text list "msjOp0": 20 'Alarma produs aparut anormal Confirmati prezenta ,integritatea si pozitia produs(planeitate , incadrarea in margini).'; 10 'Alarma detectie produs pierduta Verificati daca produsul mai exista in statie'; 11 'Alarma detectie produs pierduta Produsul exista dar nu e detectat. Reparati/ajustati senzorul de prezenta ssssssssssssssss,astfel incat sa detecteze produsul.'; 21 'Alarma produs aparut anormal Produsul nu a fost confirmat de operator Reparati senzorul ca sa nu mai indice prezenta produs'; 30 'Produsul nu a ajuns de la primul punct la al 2 lea Confirmati unde e de fapt produsul.'; 70 'Aduceti cilindru cccccccccccccc in pozitia xxxxxxxxxxxxxxx'; 72 'Deoarece a fost o alarma de griper confirmati prezenta ,integritatea si pozitia produs(planeitate , incadrarea in margini) in griper cccccccccccccc si lipsa lui de pe conveyor'; 73 'Deoarece a fost o alarma de griper confirmati prezenta ,integritatea si pozitia produs(planeitate , incadrarea in margini) pe palet si lipsa lui din griper cccccccccccccccccc'; 74 'Deoarece a fost o eroare de cilindru,confirmati ca liftul e sus si pachetul asezat pe el'; 71 ''; 22 'Alarma produs aparut anormal Produsul nu e asezat corect. Deschideti usa si plasati corect sau evacuati manual produsul,apoi validati'; 12 'Alarma detectie produs pierduta Produsul exista dar e prost asezat Deschideti usa si asezati sau eliminati produsul ,apoi confirmati.'; 31 'Produsul nu a ajuns de la primul punct la al 2 lea Produsul exista la destinatie dar nu e detectat.Deschideti usa si asezati produsul in dreptul senzorului ,sau reparati senzorul astfel incat sa detecteze produsul'; 32 'Produsul nu a ajuns de la primul punct la al 2 lea Produsul a ajuns la destinatie . Verificati prezenta,integritatea si pozitia lui si confirmati .'; 33 'Produsul nu a ajuns de la primul punct la al 2 lea Produsul a disparut din zona in mod necontrolat .Confirmati ca nici un produs nu se gaseste intre cele 2 posturi ,pentru a declara zona goala, si a putea accepta alte produse.'; 13 'Alarma detectie produs pierduta Detectia produsului a revenit Confirmati existenta si pozitia produs.'; 23 'Alarma produs aparut anormal Detectia produsului a disparut. Confirmati daca produsul mai exista'; 75 ''; 14 'Alarma detectie produs pierduta Produsul nu exista dar e detectat. Reparati/ajustati senzorul de prezenta ,astfel incat sa nu detecteze produsul.'

text list "numeOp": 0 'Conveyor intrare'; 1 'Lift intrare jos'; 2 'Lift impingator'; 3 'Conveyor iesire poz1'; 4 'Conveyor iesire poz2'; 5 'Griper robot poz 1'; 6 'Griper robot poz 2'; 7 'Impingator lift'

text list "ButOp1": 10 'Produs exista si e conform'; 11 'Produs exista si e conform'; 12 'Produs exista si e conform'; 13 'Produs exista si e conform'; 20 'Produs exista si e conform'; 21 'Produs exista si e conform'; 22 'Produs exista si e conform'; 23 'Produs exista si e conform'; 30 'Produs existala destinatie'; 31 'Produs existala destinatie'; 32 'Produs existala destinatie'; 33 'Produs existala destinatie'

text list "loc1": 1 'Locatie'; 2 'Locatie'; 3 'Plecare'

text list "ButOp2": 10 'Produs NU exista'; 11 'Produs NU exista'; 12 'Produs NU exista'; 13 'Produs NU exista'; 20 'Produs NU exista'; 21 'Produs NU exista'; 22 'Produs NU exista'; 23 'Produs NU exista'; 30 'Produs NU exista de la sursa pana la destinatie'; 31 'Produs NU exista de la sursa pana la destinatie'; 32 'Produs NU exista de la sursa pana la destinatie'; 33 'Produs NU exista de la sursa pana la destinatie'

text list "ButOp3": 10 'Produs exista dar e prost asezat'; 11 'Produs exista dar e prost asezat'; 12 'Produs exista dar e prost asezat'; 13 'Produs exista dar e prost asezat'; 20 'Produs exista dar e prost asezat'; 21 'Produs exista dar e prost asezat'; 22 'Produs exista dar e prost asezat'; 23 'Produs exista dar e prost asezat'; 30 'Produs exista linainte de destinatie'; 31 'Produs exista linainte de destinatie'; 32 'Produs exista linainte de destinatie'; 33 'Produs exista linainte de destinatie'

text list "loc2": 0..2 ''; 3 'Sosire'

graphic list "@DiagnosticsStates": 0 '@Diagnostics_StateGood'; 1 '@Diagnostics_StateBad'

screen "Alarms" 800x480, template "TemplateWithClockAndBackBtn"
   AlarmView "Alarm view_1" at 0,40 size 800x348
   Button "Button_1" at 648,392 size 144x80; TextOff 'Confirmare Alarma Acknowledge'; Authorization "Operate"
      on Press: function_d9204949("Alarm view_1"); function_b14e0dd5("DB20_DATA_HMI_Reset_Faults", 0)
   Button "Button_2" at 8,392 size 144x80; TextOff 'Loguri Sistem / Acknowledge'; Authorization "Operate"
      on Press: ActivateScreen("SystemHealth", 0)

screen "SystemHealth" 800x480, template "TemplateWithClockAndBackBtn"
   SysDiagControl "System diagnostics view_1" at 0,40 size 800x440

screen "Settings" 800x480, template "TemplateWithClockAndBackBtn"
   UserView "User view_1" at 8,48 size 784x328
   Button "Button_1" at 8,392 size 96x80; TextOff 'Reset General'; Authorization "Operate"
   Button "Button_2" at 112,392 size 96x80; TextOff 'Reset Contoare'; Authorization "Operate"
   Button "Button_3" at 216,392 size 96x80; TextOff 'Calibrare Ecran'; Authorization "Operate"
      on Press: function_bc3e350c()
   Button "Button_4" at 320,392 size 96x80; TextOff 'Curatare Ecran'; Authorization "Operate"
      on Press: function_be740847(30)
   Button "Button_5" at 424,392 size 96x80; TextOff 'Stop Runtime'; Authorization "Operate"
      on Press: StopRuntime(0)

screen "Production.Repair" 800x480, template "TemplateWithClockAndBackBtnForStatistics"
   IOField "I/O field_1" at 696,48 size 96x32; FormatPattern 9
      ProcessValue <- "PalletsLastWeek"
   TextField "Text field_1" at 488,48 size 160x20; Text 'Paleti ultima saptamana'
   TextField "Text field_2" at 488,88 size 115x20; Text 'Paleti ultima luna'
   IOField "I/O field_2" at 696,88 size 96x32; FormatPattern 9
      ProcessValue <- "PalletsLastMonth"
   TrendView "Trend view_1" at 8,48 size 448x332
   IOField "I/O field_3" at 696,127 size 96x32; FormatPattern 99
      ProcessValue <- "DB20_DATA_HMI_Step_Destacker"
   TextField "Text field_3" at 488,127 size 97x20; Text 'Pas destivuire'
   TextField "Text field_4" at 488,167 size 81x20; Text 'Pas stivuire'
   IOField "I/O field_4" at 696,167 size 96x32; FormatPattern 99
      ProcessValue <- "DB20_DATA_HMI_Step_Stacker"
   Button "Button_1" at 488,256 size 124x97; TextOff 'REZ G7 DS'
      on Release: ResetBit("Rez_G7_DS")
      on Press: SetBit("Rez_G7_DS")
   Button "Button_2" at 650,256 size 124x97; TextOff 'REZ G7 S'
      on Release: ResetBit("Rez_G7_S")
      on Press: SetBit("Rez_G7_S")

screen "Production.Destroy" 800x480, template "TemplateWithClockAndBackBtnForStatistics"
   TrendView "Trend view_1" at 8,48 size 448x332

screen "Energy" 800x480, template "TemplateWithClockAndBackBtnForStatistics"
   IOField "I/O field_1" at 688,48 size 96x32; FormatPattern 9
      ProcessValue <- "FB_EnergyCounter_DB_Counters_LastHour_CV"
   TextField "Text field_3" at 600,48 size 70x20; Text 'Ultima ora'
   IOField "I/O field_2" at 688,88 size 96x32; FormatPattern 9
      ProcessValue <- "FB_EnergyCounter_DB_Counters_LastDay_CV"
   TextField "Text field_1" at 600,88 size 58x20; Text 'Ultima zi'
   IOField "I/O field_3" at 688,128 size 96x32; FormatPattern 9
      ProcessValue <- "FB_EnergyCounter_DB_Counters_LastMonth_CV"
   TextField "Text field_2" at 600,128 size 75x20; Text 'Ultima luna'
   TrendView "Trend view_1" at 8,48 size 448x332

screen "Safety" 800x480, template "TemplateWithClockAndBackBtnForStatistics"
   IOField "I/O field_1" at 336,48 size 96x32; FormatPattern 9
      ProcessValue <- "FB_AlarmCounter_DB_Counters_Destacker 110KF1 Safety Relay_CV"
   TextField "Text field_3" at 16,50 size 208x20; Text 'Destacker 110KF1 Safety Relay'
   IOField "I/O field_2" at 336,80 size 96x32; FormatPattern 9
      ProcessValue <- "FB_AlarmCounter_DB_Counters_Destacker 111KF1 Safety Barrier Relay_CV"
   TextField "Text field_1" at 16,82 size 257x20; Text 'Destacker 111KF1 Safety Barrier Relay'
   IOField "I/O field_3" at 336,112 size 96x32; FormatPattern 9
      ProcessValue <- "FB_AlarmCounter_DB_Counters_Zone 2 112KF1 Safety Relay_CV"
   TextField "Text field_2" at 16,114 size 185x20; Text 'Zone 2 112KF1 Safety Relay'
   IOField "I/O field_4" at 336,144 size 96x32; FormatPattern 9
      ProcessValue <- "FB_AlarmCounter_DB_Counters_Stacker 113KF1 Safety Relay_CV"
   TextField "Text field_4" at 16,146 size 192x20; Text 'Stacker 113KF1 Safety Relay'
   IOField "I/O field_5" at 336,176 size 96x32; FormatPattern 9
      ProcessValue <- "FB_AlarmCounter_DB_Counters_Stacker 114KF1 Safety Barrier Relay 1_CV"
   TextField "Text field_5" at 16,178 size 253x20; Text 'Stacker 114KF1 Safety Barrier Relay 1'
   IOField "I/O field_6" at 336,208 size 96x32; FormatPattern 9
      ProcessValue <- "FB_AlarmCounter_DB_Counters_Stacker 115KF1 Safety Barrier Relay 2_CV"
   TextField "Text field_6" at 16,210 size 253x20; Text 'Stacker 115KF1 Safety Barrier Relay 2'
   IOField "I/O field_7" at 336,240 size 96x32; FormatPattern 9
      ProcessValue <- "FB_AlarmCounter_DB_Counters_Emergency Stop Destacker_CV"
   TextField "Text field_7" at 16,242 size 180x20; Text 'Emergency Stop Destacker'
   IOField "I/O field_8" at 336,272 size 96x32; FormatPattern 9
      ProcessValue <- "FB_AlarmCounter_DB_Counters_Emergency Stop Zone 2_CV"
   TextField "Text field_8" at 16,274 size 157x20; Text 'Emergency Stop Zone 2'
   IOField "I/O field_9" at 336,304 size 96x32; FormatPattern 9
      ProcessValue <- "FB_AlarmCounter_DB_Counters_Emergency Stop Stacker_CV"
   TextField "Text field_9" at 16,306 size 164x20; Text 'Emergency Stop Stacker'
   Button "Button_1" at 552,160 size 128x64; TextOff 'Reset'; Authorization "User administration"

screen "Manual.General" 800x480, template "TemplateWithClockAndBackBtnForManual"
   GraphicIOField "PlotLight_Round_G" at 224,240 size 24x24; PictureOn "PilotLight_Round_G_On_256c"; PictureOff "PilotLight_Round_G_Off_256c"
      ProcessValue <- "Prezenta aer"
   TextField "Text field_1" at 8,242 size 90x20; Text 'Prezenta aer'
   GraphicIOField "PlotLight_Round_G_1" at 224,48 size 24x24; PictureOff "PilotLight_Round_G_Off_256c"; PictureOn "PilotLight_Round_G_On_256c"
      ProcessValue <- "Aliniere palet"
   TextField "Text field_2" at 8,50 size 91x20; Text 'Aliniere palet'
   GraphicIOField "PlotLight_Round_G_2" at 224,80 size 24x24; PictureOn "PilotLight_Round_G_On_256c"; PictureOff "PilotLight_Round_G_Off_256c"
      ProcessValue <- "Centror extins"
   TextField "Text field_3" at 8,82 size 98x20; Text 'Centror extins'
   GraphicIOField "PlotLight_Round_G_3" at 224,112 size 24x24; PictureOn "PilotLight_Round_G_On_256c"; PictureOff "PilotLight_Round_G_Off_256c"
      ProcessValue <- "Centror retras"
   TextField "Text field_4" at 8,114 size 100x20; Text 'Centror retras'
   GraphicIOField "PlotLight_Round_G_6" at 224,144 size 24x24; PictureOn "PilotLight_Round_G_On_256c"; PictureOff "PilotLight_Round_G_Off_256c"
      ProcessValue <- "Detectie palet"
   TextField "Text field_7" at 8,146 size 97x20; Text 'Detectie palet'
   GraphicIOField "PlotLight_Round_G_7" at 224,176 size 24x24; PictureOff "PilotLight_Round_G_Off_256c"; PictureOn "PilotLight_Round_G_On_256c"
      ProcessValue <- "Feed palet"
   TextField "Text field_8" at 8,178 size 72x20; Text 'Feed palet'
   GraphicIOField "PlotLight_Round_G_9" at 224,208 size 24x24; PictureOff "PilotLight_Round_G_Off_256c"; PictureOn "PilotLight_Round_G_On_256c"
      ProcessValue <- "Masurare lungime"
   TextField "Text field_10" at 8,210 size 120x20; Text 'Masurare lungime'
   GraphicIOField "PlotLight_Round_G_10" at 224,272 size 24x24; PictureOff "PilotLight_Round_G_Off_256c"; PictureOn "PilotLight_Round_G_On_256c"
      ProcessValue <- "Prezenta palet iesire"
   TextField "Text field_11" at 8,274 size 140x20; Text 'Prezenta palet iesire'
   GraphicIOField "PlotLight_Round_G_11" at 224,304 size 24x24; PictureOff "PilotLight_Round_G_Off_256c"; PictureOn "PilotLight_Round_G_On_256c"
      ProcessValue <- "Prezenta palet_capat_conveyor"
   TextField "Text field_12" at 8,306 size 215x20; Text 'Prezenta palet_capat_conveyor'
   GraphicIOField "PlotLight_Round_G_12" at 224,336 size 24x24; PictureOff "PilotLight_Round_G_Off_256c"; PictureOn "PilotLight_Round_G_On_256c"
      ProcessValue <- "Prezenta palet_centror"
   TextField "Text field_13" at 8,338 size 158x20; Text 'Prezenta palet_centror'
   GraphicIOField "PlotLight_Round_G_14" at 504,264 size 24x24; PictureOff "PilotLight_Round_G_Off_256c"; PictureOn "PilotLight_Round_G_On_256c"
      ProcessValue <- "Protectie cuplata Post reparatii minore"
   TextField "Text field_15" at 264,266 size 230x20; Text 'Prot. cuplata Post reparatii minore'
   GraphicIOField "PlotLight_Round_G_15" at 504,48 size 24x24; PictureOn "PilotLight_Round_G_On_256c"; PictureOff "PilotLight_Round_G_Off_256c"
      ProcessValue <- "Prezenta palet_stanga"
   TextField "Text field_16" at 264,50 size 154x20; Text 'Prezenta palet_stanga'
   GraphicIOField "PlotLight_Round_G_16" at 504,72 size 24x24; PictureOff "PilotLight_Round_G_Off_256c"; PictureOn "PilotLight_Round_G_On_256c"
      ProcessValue <- "Prezenta stiva"
   TextField "Text field_17" at 264,74 size 100x20; Text 'Prezenta stiva'
   GraphicIOField "PlotLight_Round_G_17" at 504,96 size 24x24; PictureOff "PilotLight_Round_G_Off_256c"; PictureOn "PilotLight_Round_G_On_256c"
      ProcessValue <- "Prezenta_stiva"
   TextField "Text field_18" at 264,98 size 104x20; Text 'Prezenta_stiva'
   GraphicIOField "PlotLight_Round_G_18" at 504,120 size 24x24; PictureOff "PilotLight_Round_G_Off_256c"; PictureOn "PilotLight_Round_G_On_256c"
      ProcessValue <- "Protectie cuplata Circular masa fixa"
   TextField "Text field_19" at 264,122 size 235x20; Text 'Protectie cuplata Circular masa fixa'
   GraphicIOField "PlotLight_Round_G_19" at 504,144 size 24x24; PictureOff "PilotLight_Round_G_Off_256c"; PictureOn "PilotLight_Round_G_On_256c"
      ProcessValue <- "Protectie cuplata HMI"
   TextField "Text field_20" at 264,146 size 146x20; Text 'Protectie cuplata HMI'
   GraphicIOField "PlotLight_Round_G_20" at 504,168 size 24x24; PictureOff "PilotLight_Round_G_Off_256c"; PictureOn "PilotLight_Round_G_On_256c"
      ProcessValue <- "Protectie cuplata Iluminat"
   TextField "Text field_21" at 264,170 size 173x20; Text 'Protectie cuplata Iluminat'
   GraphicIOField "PlotLight_Round_G_21" at 504,192 size 24x24; PictureOn "PilotLight_Round_G_On_256c"; PictureOff "PilotLight_Round_G_Off_256c"
      ProcessValue <- "Protectie cuplata Masina demontare paleti dreapta"
   TextField "Text field_22" at 264,194 size 241x20; Text 'Prot. cuplata Mas. dem. pal. dreapta'
   GraphicIOField "PlotLight_Round_G_22" at 504,216 size 24x24; PictureOn "PilotLight_Round_G_On_256c"; PictureOff "PilotLight_Round_G_Off_256c"
      ProcessValue <- "Protectie cuplata Masina demontare paleti stanga"
   TextField "Text field_23" at 264,218 size 234x20; Text 'Prot. cuplata Mas. dem. pal. stanga'
   GraphicIOField "PlotLight_Round_G_23" at 504,240 size 24x24; PictureOn "PilotLight_Round_G_On_256c"; PictureOff "PilotLight_Round_G_Off_256c"
      ProcessValue <- "Protectie cuplata Post reparatie stanga+dreapta"
   TextField "Text field_24" at 264,242 size 218x20; Text 'Prot. cuplata Post rep. stg.+drp.'
   GraphicIOField "PlotLight_Round_G_24" at 504,288 size 24x24; PictureOn "PilotLight_Round_G_On_256c"; PictureOff "PilotLight_Round_G_Off_256c"
      ProcessValue <- "Protectie cuplata TELE"
   TextField "Text field_25" at 264,290 size 149x20; Text 'Protectie cuplata TELE'
   GraphicIOField "PlotLight_Round_G_25" at 504,312 size 24x24; PictureOn "PilotLight_Round_G_On_256c"; PictureOff "PilotLight_Round_G_Off_256c"
      ProcessValue <- "Prezenta palet_capat_conveyor"
   TextField "Text field_26" at 264,314 size 215x20; Text 'Prezenta palet_capat_conveyor'
   GraphicIOField "PlotLight_Round_G_26" at 504,336 size 24x24; PictureOn "PilotLight_Round_G_On_256c"; PictureOff "PilotLight_Round_G_Off_256c"
      ProcessValue <- "Prezenta palet_centror"
   TextField "Text field_27" at 264,338 size 158x20; Text 'Prezenta palet_centror'
   GraphicIOField "PlotLight_Round_G_31" at 760,48 size 24x24; PictureOn "PilotLight_Round_G_On_256c"; PictureOff "PilotLight_Round_G_Off_256c"
      ProcessValue <- "Senzor 1 proximitate softstarter aer zona 2"
   TextField "Text field_32" at 544,50 size 206x20; Text 'Senzor 1 prox. soft. aer zona 2'
   GraphicIOField "PlotLight_Round_G_35" at 760,84 size 24x24; PictureOn "PilotLight_Round_G_On_256c"; PictureOff "PilotLight_Round_G_Off_256c"
      ProcessValue <- "Senzor 2 proximitate softstarter aer zona 2"
   TextField "Text field_36" at 544,86 size 206x20; Text 'Senzor 2 prox. soft. aer zona 2'
   GraphicIOField "PlotLight_Round_G_36" at 760,120 size 24x24; PictureOn "PilotLight_Round_G_On_256c"; PictureOff "PilotLight_Round_G_Off_256c"
      ProcessValue <- "Senzor destacking"
   TextField "Text field_37" at 544,122 size 124x20; Text 'Senzor destacking'
   GraphicIOField "PlotLight_Round_G_37" at 760,156 size 24x24; PictureOff "PilotLight_Round_G_Off_256c"; PictureOn "PilotLight_Round_G_On_256c"
      ProcessValue <- "Senzor stacking"
   TextField "Text field_38" at 544,158 size 108x20; Text 'Senzor stacking'
   GraphicIOField "PlotLight_Round_G_38" at 760,192 size 24x24; PictureOff "PilotLight_Round_G_Off_256c"; PictureOn "PilotLight_Round_G_On_256c"
      ProcessValue <- "Start masurare lungime"
   TextField "Text field_39" at 544,194 size 158x20; Text 'Start masurare lungime'

screen "Manual.IOLinkDiag" 800x480, template "TemplateWithClockAndBackBtnForManual"
   GraphicIOField "PlotLight_Round_G" at 136,48 size 24x24; PictureOff "PilotLight_Round_G_Off_256c"; PictureOn "PilotLight_Round_G_On_256c"
      ProcessValue <- "MD_IS1_SC_X1.0"
   TextField "Text field_1" at 8,50 size 115x20; Text 'MD_IS1_SC_X1.0'
   GraphicIOField "PlotLight_Round_G_1" at 136,72 size 24x24; PictureOn "PilotLight_Round_G_On_256c"; PictureOff "PilotLight_Round_G_Off_256c"
      ProcessValue <- "MD_IS1_SC_X1.1"
   TextField "Text field_2" at 8,74 size 115x20; Text 'MD_IS1_SC_X1.1'
   GraphicIOField "PlotLight_Round_G_2" at 136,96 size 24x24; PictureOn "PilotLight_Round_G_On_256c"; PictureOff "PilotLight_Round_G_Off_256c"
      ProcessValue <- "MD_IS1_SC_X1.2"
   TextField "Text field_3" at 8,98 size 115x20; Text 'MD_IS1_SC_X1.2'
   GraphicIOField "PlotLight_Round_G_3" at 136,120 size 24x24; PictureOff "PilotLight_Round_G_Off_256c"; PictureOn "PilotLight_Round_G_On_256c"
      ProcessValue <- "MD_IS1_SC_X1.3"
   TextField "Text field_4" at 8,122 size 115x20; Text 'MD_IS1_SC_X1.3'
   GraphicIOField "PlotLight_Round_G_4" at 136,144 size 24x24; PictureOff "PilotLight_Round_G_Off_256c"; PictureOn "PilotLight_Round_G_On_256c"
      ProcessValue <- "MD_IS1_SC_X1.4"
   TextField "Text field_5" at 8,146 size 115x20; Text 'MD_IS1_SC_X1.4'
   GraphicIOField "PlotLight_Round_G_5" at 136,168 size 24x24; PictureOff "PilotLight_Round_G_Off_256c"; PictureOn "PilotLight_Round_G_On_256c"
      ProcessValue <- "MD_IS1_SC_X1.5"
   TextField "Text field_6" at 8,170 size 115x20; Text 'MD_IS1_SC_X1.5'
   GraphicIOField "PlotLight_Round_G_6" at 136,192 size 24x24; PictureOff "PilotLight_Round_G_Off_256c"; PictureOn "PilotLight_Round_G_On_256c"
      ProcessValue <- "MD_IS1_SC_X1.6"
   TextField "Text field_7" at 8,194 size 115x20; Text 'MD_IS1_SC_X1.6'
   GraphicIOField "PlotLight_Round_G_7" at 136,216 size 24x24; PictureOff "PilotLight_Round_G_Off_256c"; PictureOn "PilotLight_Round_G_On_256c"
      ProcessValue <- "MD_IS1_SC_X1.7"
   TextField "Text field_8" at 8,218 size 115x20; Text 'MD_IS1_SC_X1.7'
   GraphicIOField "PlotLight_Round_G_8" at 312,48 size 24x24; PictureOn "PilotLight_Round_G_On_256c"; PictureOff "PilotLight_Round_G_Off_256c"
      ProcessValue <- "MD_IS2_SC_X1.0"
   TextField "Text field_9" at 184,50 size 115x20; Text 'MD_IS2_SC_X1.0'
   GraphicIOField "PlotLight_Round_G_9" at 312,72 size 24x24; PictureOff "PilotLight_Round_G_Off_256c"; PictureOn "PilotLight_Round_G_On_256c"
      ProcessValue <- "MD_IS2_SC_X1.1"
   TextField "Text field_10" at 184,74 size 115x20; Text 'MD_IS2_SC_X1.1'
   GraphicIOField "PlotLight_Round_G_10" at 312,96 size 24x24; PictureOff "PilotLight_Round_G_Off_256c"; PictureOn "PilotLight_Round_G_On_256c"
      ProcessValue <- "MD_IS2_SC_X1.2"
   TextField "Text field_11" at 184,98 size 115x20; Text 'MD_IS2_SC_X1.2'
   GraphicIOField "PlotLight_Round_G_11" at 312,120 size 24x24; PictureOn "PilotLight_Round_G_On_256c"; PictureOff "PilotLight_Round_G_Off_256c"
      ProcessValue <- "MD_IS2_SC_X1.3"
   TextField "Text field_12" at 184,122 size 115x20; Text 'MD_IS2_SC_X1.3'
   GraphicIOField "PlotLight_Round_G_12" at 312,144 size 24x24; PictureOn "PilotLight_Round_G_On_256c"; PictureOff "PilotLight_Round_G_Off_256c"
      ProcessValue <- "MD_IS2_SC_X1.4"
   TextField "Text field_13" at 184,146 size 115x20; Text 'MD_IS2_SC_X1.4'
   GraphicIOField "PlotLight_Round_G_13" at 312,168 size 24x24; PictureOn "PilotLight_Round_G_On_256c"; PictureOff "PilotLight_Round_G_Off_256c"
      ProcessValue <- "MD_IS2_SC_X1.5"
   TextField "Text field_14" at 184,170 size 115x20; Text 'MD_IS2_SC_X1.5'
   GraphicIOField "PlotLight_Round_G_14" at 312,192 size 24x24; PictureOn "PilotLight_Round_G_On_256c"; PictureOff "PilotLight_Round_G_Off_256c"
      ProcessValue <- "MD_IS2_SC_X1.6"
   TextField "Text field_15" at 184,194 size 115x20; Text 'MD_IS2_SC_X1.6'
   GraphicIOField "PlotLight_Round_G_15" at 312,216 size 24x24; PictureOn "PilotLight_Round_G_On_256c"; PictureOff "PilotLight_Round_G_Off_256c"
      ProcessValue <- "MD_IS2_SC_X1.7"
   TextField "Text field_16" at 184,218 size 115x20; Text 'MD_IS2_SC_X1.7'
   GraphicIOField "PlotLight_Round_G_16" at 136,240 size 24x24; PictureOff "PilotLight_Round_G_Off_256c"; PictureOn "PilotLight_Round_G_On_256c"
      ProcessValue <- "MD_OS_SC_X1.0"
   TextField "Text field_17" at 8,242 size 111x20; Text 'MD_OS_SC_X1.0'
   GraphicIOField "PlotLight_Round_G_17" at 136,264 size 24x24; PictureOn "PilotLight_Round_G_On_256c"; PictureOff "PilotLight_Round_G_Off_256c"
      ProcessValue <- "MD_OS_SC_X1.1"
   TextField "Text field_18" at 8,266 size 111x20; Text 'MD_OS_SC_X1.1'
   GraphicIOField "PlotLight_Round_G_18" at 136,288 size 24x24; PictureOn "PilotLight_Round_G_On_256c"; PictureOff "PilotLight_Round_G_Off_256c"
      ProcessValue <- "MD_OS_SC_X1.2"
   TextField "Text field_19" at 8,290 size 111x20; Text 'MD_OS_SC_X1.2'
   GraphicIOField "PlotLight_Round_G_19" at 136,312 size 24x24; PictureOff "PilotLight_Round_G_Off_256c"; PictureOn "PilotLight_Round_G_On_256c"
      ProcessValue <- "MD_OS_SC_X1.3"
   TextField "Text field_20" at 8,314 size 111x20; Text 'MD_OS_SC_X1.3'
   GraphicIOField "PlotLight_Round_G_20" at 136,336 size 24x24; PictureOff "PilotLight_Round_G_Off_256c"; PictureOn "PilotLight_Round_G_On_256c"
      ProcessValue <- "MD_OS_SC_X1.4"
   TextField "Text field_21" at 8,338 size 111x20; Text 'MD_OS_SC_X1.4'
   GraphicIOField "PlotLight_Round_G_21" at 136,360 size 24x24; PictureOff "PilotLight_Round_G_Off_256c"; PictureOn "PilotLight_Round_G_On_256c"
      ProcessValue <- "MD_OS_SC_X1.5"
   TextField "Text field_22" at 8,362 size 111x20; Text 'MD_OS_SC_X1.5'
   GraphicIOField "PlotLight_Round_G_22" at 488,48 size 24x24; PictureOn "PilotLight_Round_G_On_256c"; PictureOff "PilotLight_Round_G_Off_256c"
      ProcessValue <- "MS_IS1_SC_X1.0"
   TextField "Text field_23" at 360,50 size 114x20; Text 'MS_IS1_SC_X1.0'
   GraphicIOField "PlotLight_Round_G_23" at 488,72 size 24x24; PictureOff "PilotLight_Round_G_Off_256c"; PictureOn "PilotLight_Round_G_On_256c"
      ProcessValue <- "MS_IS1_SC_X1.1"
   TextField "Text field_24" at 360,74 size 114x20; Text 'MS_IS1_SC_X1.1'
   GraphicIOField "PlotLight_Round_G_24" at 488,96 size 24x24; PictureOff "PilotLight_Round_G_Off_256c"; PictureOn "PilotLight_Round_G_On_256c"
      ProcessValue <- "MS_IS1_SC_X1.2"
   TextField "Text field_25" at 360,98 size 114x20; Text 'MS_IS1_SC_X1.2'
   GraphicIOField "PlotLight_Round_G_25" at 488,120 size 24x24; PictureOn "PilotLight_Round_G_On_256c"; PictureOff "PilotLight_Round_G_Off_256c"
      ProcessValue <- "MS_IS1_SC_X1.3"
   TextField "Text field_26" at 360,122 size 114x20; Text 'MS_IS1_SC_X1.3'
   GraphicIOField "PlotLight_Round_G_26" at 488,144 size 24x24; PictureOn "PilotLight_Round_G_On_256c"; PictureOff "PilotLight_Round_G_Off_256c"
      ProcessValue <- "MS_IS1_SC_X1.4"
   TextField "Text field_27" at 360,146 size 114x20; Text 'MS_IS1_SC_X1.4'
   GraphicIOField "PlotLight_Round_G_27" at 488,168 size 24x24; PictureOn "PilotLight_Round_G_On_256c"; PictureOff "PilotLight_Round_G_Off_256c"
      ProcessValue <- "MS_IS1_SC_X1.5"
   TextField "Text field_28" at 360,170 size 114x20; Text 'MS_IS1_SC_X1.5'
   GraphicIOField "PlotLight_Round_G_28" at 488,192 size 24x24; PictureOn "PilotLight_Round_G_On_256c"; PictureOff "PilotLight_Round_G_Off_256c"
      ProcessValue <- "MS_IS1_SC_X1.6"
   TextField "Text field_29" at 360,194 size 114x20; Text 'MS_IS1_SC_X1.6'
   GraphicIOField "PlotLight_Round_G_29" at 488,216 size 24x24; PictureOn "PilotLight_Round_G_On_256c"; PictureOff "PilotLight_Round_G_Off_256c"
      ProcessValue <- "MS_IS1_SC_X1.7"
   TextField "Text field_30" at 360,218 size 114x20; Text 'MS_IS1_SC_X1.7'
   GraphicIOField "PlotLight_Round_G_30" at 664,48 size 24x24; PictureOff "PilotLight_Round_G_Off_256c"; PictureOn "PilotLight_Round_G_On_256c"
      ProcessValue <- "MS_IS2_SC_X1.0"
   TextField "Text field_31" at 536,50 size 114x20; Text 'MS_IS2_SC_X1.0'
   GraphicIOField "PlotLight_Round_G_31" at 664,72 size 24x24; PictureOn "PilotLight_Round_G_On_256c"; PictureOff "PilotLight_Round_G_Off_256c"
      ProcessValue <- "MS_IS2_SC_X1.1"
   TextField "Text field_32" at 536,74 size 114x20; Text 'MS_IS2_SC_X1.1'
   GraphicIOField "PlotLight_Round_G_32" at 664,96 size 24x24; PictureOn "PilotLight_Round_G_On_256c"; PictureOff "PilotLight_Round_G_Off_256c"
      ProcessValue <- "MS_IS2_SC_X1.2"
   TextField "Text field_33" at 536,98 size 114x20; Text 'MS_IS2_SC_X1.2'
   GraphicIOField "PlotLight_Round_G_33" at 664,120 size 24x24; PictureOff "PilotLight_Round_G_Off_256c"; PictureOn "PilotLight_Round_G_On_256c"
      ProcessValue <- "MS_IS2_SC_X1.3"
   TextField "Text field_34" at 536,122 size 114x20; Text 'MS_IS2_SC_X1.3'
   GraphicIOField "PlotLight_Round_G_34" at 664,144 size 24x24; PictureOff "PilotLight_Round_G_Off_256c"; PictureOn "PilotLight_Round_G_On_256c"
      ProcessValue <- "MS_IS2_SC_X1.4"
   TextField "Text field_35" at 536,146 size 114x20; Text 'MS_IS2_SC_X1.4'
   GraphicIOField "PlotLight_Round_G_35" at 664,168 size 24x24; PictureOff "PilotLight_Round_G_Off_256c"; PictureOn "PilotLight_Round_G_On_256c"
      ProcessValue <- "MS_IS2_SC_X1.5"
   TextField "Text field_36" at 536,170 size 114x20; Text 'MS_IS2_SC_X1.5'
   GraphicIOField "PlotLight_Round_G_36" at 664,192 size 24x24; PictureOff "PilotLight_Round_G_Off_256c"; PictureOn "PilotLight_Round_G_On_256c"
      ProcessValue <- "MS_IS2_SC_X1.6"
   TextField "Text field_37" at 536,194 size 114x20; Text 'MS_IS2_SC_X1.6'
   GraphicIOField "PlotLight_Round_G_37" at 664,216 size 24x24; PictureOff "PilotLight_Round_G_Off_256c"; PictureOn "PilotLight_Round_G_On_256c"
      ProcessValue <- "MS_IS2_SC_X1.7"
   TextField "Text field_38" at 536,218 size 114x20; Text 'MS_IS2_SC_X1.7'
   GraphicIOField "PlotLight_Round_G_38" at 488,240 size 24x24; PictureOn "PilotLight_Round_G_On_256c"; PictureOff "PilotLight_Round_G_Off_256c"
      ProcessValue <- "MS_OS_SC_X1.0"
   TextField "Text field_39" at 360,242 size 110x20; Text 'MS_OS_SC_X1.0'
   GraphicIOField "PlotLight_Round_G_39" at 488,264 size 24x24; PictureOff "PilotLight_Round_G_Off_256c"; PictureOn "PilotLight_Round_G_On_256c"
      ProcessValue <- "MS_OS_SC_X1.1"
   TextField "Text field_40" at 360,266 size 110x20; Text 'MS_OS_SC_X1.1'
   GraphicIOField "PlotLight_Round_G_40" at 488,288 size 24x24; PictureOff "PilotLight_Round_G_Off_256c"; PictureOn "PilotLight_Round_G_On_256c"
      ProcessValue <- "MS_OS_SC_X1.2"
   TextField "Text field_41" at 360,290 size 110x20; Text 'MS_OS_SC_X1.2'
   GraphicIOField "PlotLight_Round_G_41" at 488,312 size 24x24; PictureOn "PilotLight_Round_G_On_256c"; PictureOff "PilotLight_Round_G_Off_256c"
      ProcessValue <- "MS_OS_SC_X1.3"
   TextField "Text field_42" at 360,314 size 110x20; Text 'MS_OS_SC_X1.3'
   GraphicIOField "PlotLight_Round_G_42" at 488,336 size 24x24; PictureOn "PilotLight_Round_G_On_256c"; PictureOff "PilotLight_Round_G_Off_256c"
      ProcessValue <- "MS_OS_SC_X1.4"
   TextField "Text field_43" at 360,338 size 110x20; Text 'MS_OS_SC_X1.4'
   GraphicIOField "PlotLight_Round_G_43" at 488,360 size 24x24; PictureOn "PilotLight_Round_G_On_256c"; PictureOff "PilotLight_Round_G_Off_256c"
      ProcessValue <- "MS_OS_SC_X1.5"
   TextField "Text field_44" at 360,362 size 110x20; Text 'MS_OS_SC_X1.5'

screen "Manual.StackerAConveyors" 800x480, template "TemplateWithClockAndBackBtnForManual"
   TextField "Text field_15" at 368,54 size 300x20; Text 'Cuplare contactor VFD Conveior 4 descarcare'
   TextField "Text field_16" at 368,94 size 297x20; Text 'Fault Aknowledge VFD Conveior 4 descarcare'
   TextField "Text field_17" at 368,134 size 237x20; Text 'ON/OFF1 VFD Conveior 4 descarcare'
   Switch "Switch_1" at 696,48 size 73x32; CaptionText 'Switch'; TextOff 'OFF'; TextOn 'ON'
      on SwitchOff: ResetBit("Manual_Cuplare contactor VFD Conveior 4 descarcare stacker")
      on SwitchOn: SetBit("Manual_Cuplare contactor VFD Conveior 4 descarcare stacker")
      ProcessValue <- "Cuplare contactor VFD Conveior 4 descarcare stacker"
   GraphicIOField "PlotLight_Round_G_2" at 288,48 size 24x24; PictureOn "PilotLight_Round_G_On_256c"; PictureOff "PilotLight_Round_G_Off_256c"
      ProcessValue <- "Avarie Conveior 4 stacker"
   TextField "Text field_3" at 16,50 size 174x20; Text 'Avarie Conveior 4 stacker'
   GraphicIOField "PlotLight_Round_G_4" at 288,72 size 24x24; PictureOn "PilotLight_Round_G_On_256c"; PictureOff "PilotLight_Round_G_Off_256c"
      ProcessValue <- "Contactor cuplat Conveior 4 descarcare stacker"
   TextField "Text field_5" at 16,74 size 264x20; Text 'Contactor cuplat Conveior 4 descarcare'
   GraphicIOField "PlotLight_Round_G_6" at 288,120 size 24x24; PictureOn "PilotLight_Round_G_On_256c"; PictureOff "PilotLight_Round_G_Off_256c"
      ProcessValue <- "Frana decuplata Conveior 4 descarcare stacker"
   TextField "Text field_7" at 16,122 size 259x20; Text 'Frana decuplata Conveior 4 descarcare'
   GraphicIOField "PlotLight_Round_G_8" at 288,96 size 24x24; PictureOn "PilotLight_Round_G_On_256c"; PictureOff "PilotLight_Round_G_Off_256c"
      ProcessValue <- "Emergency Stop Stacker"
   TextField "Text field_9" at 16,98 size 164x20; Text 'Emergency Stop Stacker'
   GraphicIOField "PlotLight_Round_G_11" at 288,144 size 24x24; PictureOn "PilotLight_Round_G_On_256c"; PictureOff "PilotLight_Round_G_Off_256c"
      ProcessValue <- "Functionare Conveior 4 stacker"
   TextField "Text field_12" at 16,146 size 207x20; Text 'Functionare Conveior 4 stacker'
   GraphicIOField "PlotLight_Round_G_1" at 288,168 size 24x24; PictureOff "PilotLight_Round_G_Off_256c"; PictureOn "PilotLight_Round_G_On_256c"
      ProcessValue <- "Protectie cuplata Conveior 4 descarcare stacker"
   TextField "Text field_1" at 16,170 size 267x20; Text 'Protectie cuplata Conveior 4 descarcare'
   Button "DS_ACK_VFD1" at 696,90 size 73x32; TextOn 'ON'; TextOff 'OFF'
      on Release: ResetBit("Manual_Fault Aknowledge VFD Conveior 4 descarcare stacker")
      on Press: SetBit("Manual_Fault Aknowledge VFD Conveior 4 descarcare stacker")
      Appearance <- "Manual_DS_Comanda cilindru vertical jos"
   Button "DS_ON/OFF_VFD1" at 696,129 size 73x32; TextOn 'ON'; TextOff 'OFF'
      on Release: ResetBit("Manual_ON/OFF1 VFD Conveior 4 descarcare stacker")
      on Press: SetBit("Manual_ON/OFF1 VFD Conveior 4 descarcare stacker")
      Appearance <- "Manual_DS_Comanda cilindru vertical jos"

screen "Manual.Safety" 800x480, template "TemplateWithClockAndBackBtnForManual"
   GraphicIOField "PlotLight_Round_G_2" at 280,48 size 24x24; PictureOn "PilotLight_Round_G_On_256c"; PictureOff "PilotLight_Round_G_Off_256c"
      ProcessValue <- "Destacker 110KF1 Safety Relay"
   TextField "Text field_3" at 16,50 size 208x20; Text 'Destacker 110KF1 Safety Relay'
   GraphicIOField "PlotLight_Round_G_1" at 280,72 size 24x24; PictureOff "PilotLight_Round_G_Off_256c"; PictureOn "PilotLight_Round_G_On_256c"
      ProcessValue <- "Destacker 111KF1 Safety Barrier Relay"
   TextField "Text field_1" at 16,74 size 257x20; Text 'Destacker 111KF1 Safety Barrier Relay'
   GraphicIOField "PlotLight_Round_G_3" at 280,96 size 24x24; PictureOn "PilotLight_Round_G_On_256c"; PictureOff "PilotLight_Round_G_Off_256c"
      ProcessValue <- "Emergency Stop Destacker"
   TextField "Text field_2" at 16,98 size 180x20; Text 'Emergency Stop Destacker'
   GraphicIOField "PlotLight_Round_G_4" at 280,120 size 24x24; PictureOff "PilotLight_Round_G_Off_256c"; PictureOn "PilotLight_Round_G_On_256c"
      ProcessValue <- "Emergency Stop Stacker"
   TextField "Text field_4" at 16,122 size 164x20; Text 'Emergency Stop Stacker'
   GraphicIOField "PlotLight_Round_G_5" at 280,144 size 24x24; PictureOff "PilotLight_Round_G_Off_256c"; PictureOn "PilotLight_Round_G_On_256c"
      ProcessValue <- "Emergency Stop Zone 2"
   TextField "Text field_5" at 16,146 size 157x20; Text 'Emergency Stop Zone 2'
   GraphicIOField "PlotLight_Round_G_6" at 280,168 size 24x24; PictureOff "PilotLight_Round_G_Off_256c"; PictureOn "PilotLight_Round_G_On_256c"
      ProcessValue <- "Stacker 113KF1 Safety Relay"
   TextField "Text field_6" at 16,170 size 192x20; Text 'Stacker 113KF1 Safety Relay'
   GraphicIOField "PlotLight_Round_G_7" at 280,192 size 24x24; PictureOff "PilotLight_Round_G_Off_256c"; PictureOn "PilotLight_Round_G_On_256c"
      ProcessValue <- "Stacker 114KF1 Safety Barrier Relay 1"
   TextField "Text field_7" at 16,194 size 253x20; Text 'Stacker 114KF1 Safety Barrier Relay 1'
   GraphicIOField "PlotLight_Round_G_8" at 280,216 size 24x24; PictureOff "PilotLight_Round_G_Off_256c"; PictureOn "PilotLight_Round_G_On_256c"
      ProcessValue <- "Stacker 115KF1 Safety Barrier Relay 2"
   TextField "Text field_8" at 16,218 size 253x20; Text 'Stacker 115KF1 Safety Barrier Relay 2'
   GraphicIOField "PlotLight_Round_G_9" at 280,240 size 24x24; PictureOff "PilotLight_Round_G_Off_256c"; PictureOn "PilotLight_Round_G_On_256c"
      ProcessValue <- "Zone 2 112KF1 Safety Relay"
   TextField "Text field_9" at 16,242 size 185x20; Text 'Zone 2 112KF1 Safety Relay'
   TextField "Text field_14" at 384,54 size 250x20; Text 'Reset Destacker 110KF1 Safety Relay'
   TextField "Text field_10" at 384,94 size 299x20; Text 'Reset Destacker 111KF1 Safety Barrier Relay'
   TextField "Text field_11" at 384,134 size 136x20; Text 'Reset safety Zone 2'
   TextField "Text field_12" at 384,174 size 234x20; Text 'Reset Stacker 113KF1 Safety Relay'
   TextField "Text field_13" at 384,214 size 295x20; Text 'Reset Stacker 114KF1 Safety Barrier Relay 1'
   TextField "Text field_15" at 384,254 size 295x20; Text 'Reset Stacker 115KF1 Safety Barrier Relay 2'
   TextField "Text field_16" at 384,294 size 227x20; Text 'Reset Zone 2 112KF1 Safety Relay'
   Button "110KF1" at 692,50 size 73x32; TextOn 'ON'; TextOff 'OFF'
      on Release: ResetBit("Manual_Reset Stacker_New 110KF1 Safety Relay")
      on Press: SetBit("Manual_Reset Stacker_New 110KF1 Safety Relay")
      Appearance <- "Manual_DS_Comanda cilindru vertical jos"
   Button "111KF1" at 692,94 size 73x32; TextOn 'ON'; TextOff 'OFF'
      on Release: ResetBit("Manual_Reset Destacker 111KF1 Safety Barrier Relay")
      on Press: SetBit("Manual_Reset Destacker 111KF1 Safety Barrier Relay")
      Appearance <- "Manual_DS_Comanda cilindru vertical jos"
   Button "112KF1" at 692,136 size 73x32; TextOn 'ON'; TextOff 'OFF'
      on Release: ResetBit("Manual_Reset Zone 2 112KF1 Safety Relay")
      on Press: SetBit("Manual_Reset Zone 2 112KF1 Safety Relay")
      Appearance <- "Manual_DS_Comanda cilindru vertical jos"
   Button "113KF1" at 692,174 size 73x32; TextOn 'ON'; TextOff 'OFF'
      on Release: ResetBit("Manual_Reset Stacker 113KF1 Safety Relay")
      on Press: SetBit("Manual_Reset Stacker 113KF1 Safety Relay")
      Appearance <- "Manual_DS_Comanda cilindru vertical jos"
   Button "114KF1" at 692,212 size 73x32; TextOn 'ON'; TextOff 'OFF'
      on Release: ResetBit("Manual_Reset Stacker 114KF1 Safety Barrier Relay 1")
      on Press: SetBit("Manual_Reset Stacker 114KF1 Safety Barrier Relay 1")
      Appearance <- "Manual_DS_Comanda cilindru vertical jos"
   Button "115KF1" at 692,250 size 73x32; TextOn 'ON'; TextOff 'OFF'
      on Release: ResetBit("Manual_Reset Stacker 115KF1 Safety Barrier Relay 2")
      on Press: SetBit("Manual_Reset Stacker 115KF1 Safety Barrier Relay 2")
      Appearance <- "Manual_DS_Comanda cilindru vertical jos"
   Button "112KF1_4" at 692,288 size 73x32; TextOn 'ON'; TextOff 'OFF'
      on Release: ResetBit("Manual_Reset Zone 2 112KF1 Safety Relay")
      on Press: SetBit("Manual_Reset Zone 2 112KF1 Safety Relay")
      Appearance <- "Manual_DS_Comanda cilindru vertical jos"